VERSION : 0.1
   VAR_INPUT
      tcon_param : TCON_Param;
      send_buffer : "ADP.Message_Buffer.UDT";
   END_VAR
   VAR_IN_OUT
      requests : "Connection_Requests.UDT";
      saved_status : "Connection_Status.UDT";
   END_VAR
   VAR
      timers : "Connection_Status_Timers.UDT";
      TSEND : TSEND;
   END_VAR
   VAR_TEMP
      block_staus : "Connection_Status.UDT";
   END_VAR
BEGIN
   #TSEND(REQ := #requests.send,
          ID := #tcon_param.ID,
          DONE => #block_staus.done,
          BUSY => #block_staus.busy,
          ERROR => #block_staus.error,
          STATUS => #block_staus.status,
          DATA := #send_buffer);
   #requests.send := FALSE;
   "Send_Status.to_Control_Element"(requests := #requests,
                                    block_status := #block_staus,
                                    saved_status := #saved_status,
                                    timers := #timers);
END_FUNCTION_BLOCK

// folder: tcpip_connection/send/send_status

FUNCTION "Send_Status.Done" : Void   // FC168, SCL
{ S7_Optimized_Access := 'TRUE' }
VERSION : 0.1
   VAR_INPUT
      requests : "Connection_Requests.UDT";
      block_status : "Connection_Status.UDT";
   END_VAR
   VAR_IN_OUT
      saved_status : "Connection_Status.UDT";
   END_VAR
BEGIN
   "Send_Status.Set_Done"(block_status := #block_status,
                                requests := #requests,
                                saved_status := #saved_status);
   "Send_Status.Reset_Done"(block_status := #block_status,
                                  requests := #requests,
                                  saved_status := #saved_status);
END_FUNCTION

FUNCTION "Send_Status.Error" : Void   // FC169, SCL
{ S7_Optimized_Access := 'TRUE' }
VERSION : 0.1
   VAR_INPUT
      block_status : "Connection_Status.UDT";
      requests : "Connection_Requests.UDT";
   END_VAR
   VAR_IN_OUT
      off_delay : TOF_TIME;
      saved_status : "Connection_Status.UDT";
   END_VAR
BEGIN
   "Send_Status.Set_Error"(block_status := #block_status,
                                 requests := #requests,
                                 off_delay := #off_delay,
                                 saved_status := #saved_status);
END_FUNCTION

FUNCTION "Send_Status.Reset_Busy" : Void   // FC170, SCL
{ S7_Optimized_Access := 'TRUE' }
VERSION : 0.1
   VAR_INPUT
      requests : "Connection_Requests.UDT";
   END_VAR
   VAR_IN_OUT
      saved_status : "Connection_Status.UDT";
   END_VAR
BEGIN
   IF #requests.connect THEN
       #saved_status.busy := FALSE;
   END_IF;
END_FUNCTION

FUNCTION "Send_Status.Set_Busy" : Void   // FC171, SCL
{ S7_Optimized_Access := 'TRUE' }
VERSION : 0.1
   VAR_INPUT
      block_status : "Connection_Status.UDT";
      requests : "Connection_Requests.UDT";
   END_VAR
   VAR_IN_OUT
      off_delay : TOF_TIME;
      saved_status : "Connection_Status.UDT";
   END_VAR
   VAR_TEMP
      _et : Time;
   END_VAR
   VAR CONSTANT
      DELAY : Time := t#3s;
   END_VAR
BEGIN
   #off_delay(IN := #block_status.busy AND NOT #requests.disconnect,
              PT := #DELAY,
              Q => #saved_status.busy,
              ET => #_et);
END_FUNCTION

FUNCTION "Send_Status.Busy" : Void   // FC172, SCL
{ S7_Optimized_Access := 'TRUE' }
VERSION : 0.1
   VAR_INPUT
      block_status : "Connection_Status.UDT";
      requests : "Connection_Requests.UDT";
   END_VAR
   VAR_IN_OUT
      off_delay : TOF_TIME;
      saved_status : "Connection_Status.UDT";
   END_VAR
BEGIN
   "Send_Status.Set_Busy"(block_status := #block_status,
                                requests := #requests,
                                off_delay := #off_delay,
                                saved_status := #saved_status);
   "Send_Status.Reset_Busy"(requests := #requests,
                                  saved_status := #saved_status);
END_FUNCTION

FUNCTION "Send_Status.to_Control_Element" : Void   // FC173, SCL
{ S7_Optimized_Access := 'TRUE' }
VERSION : 0.1
   VAR_INPUT
      requests : "Connection_Requests.UDT";
      block_status : "Connection_Status.UDT";
   END_VAR
   VAR_IN_OUT
      saved_status : "Connection_Status.UDT";
      timers : "Connection_Status_Timers.UDT";
   END_VAR
BEGIN
   "Send_Status.Busy"(block_status := #block_status,
                            requests := #requests,
                            off_delay := #timers.busy,
                            saved_status := #saved_status);
   "Send_Status.Done"(requests := #requests,
                            block_status := #block_status,
                            saved_status := #saved_status);
   "Send_Status.Error"(block_status := #block_status,
                             requests := #requests,
                             off_delay := #timers.error,
                             saved_status := #saved_status);
   "Send_Status.Status"(block_status := #block_status,
                              requests := #requests,
                              saved_status := #saved_status,
                              status_timer := #timers.status);
END_FUNCTION

FUNCTION "Send_Status.Set_Done" : Void   // FC174, SCL
{ S7_Optimized_Access := 'TRUE' }
VERSION : 0.1
   VAR_INPUT
      block_status : "Connection_Status.UDT";
      requests : "Connection_Requests.UDT";
   END_VAR
   VAR_IN_OUT
      saved_status : "Connection_Status.UDT";
   END_VAR
BEGIN
   IF #block_status.done THEN
       #saved_status.done := TRUE;
   END_IF;
END_FUNCTION

FUNCTION "Send_Status.Reset_Done" : Void   // FC175, SCL
{ S7_Optimized_Access := 'TRUE' }
VERSION : 0.1
   VAR_INPUT
      block_status : "Connection_Status.UDT";
      requests : "Connection_Requests.UDT";
   END_VAR
   VAR_IN_OUT
      saved_status : "Connection_Status.UDT";
   END_VAR
BEGIN
   IF #requests.connect THEN
       #saved_status.done := FALSE;
   END_IF;
END_FUNCTION

FUNCTION "Send_Status.Set_Error" : Void   // FC176, SCL
{ S7_Optimized_Access := 'TRUE' }
VERSION : 0.1
   VAR_INPUT
      block_status : "Connection_Status.UDT";
      requests : "Connection_Requests.UDT";
   END_VAR
   VAR_IN_OUT
      off_delay : TOF_TIME;
      saved_status : "Connection_Status.UDT";
   END_VAR
   VAR_TEMP
      _et : Time;
   END_VAR
   VAR CONSTANT
      DELAY : Time := t#30s;
   END_VAR
BEGIN
   #off_delay(IN := #block_status.error,
              PT := #DELAY,
              Q => #saved_status.error,
              ET => #_et);
END_FUNCTION

FUNCTION "Send_Status.Save_Status" : Void   // FC177, SCL
{ S7_Optimized_Access := 'TRUE' }
VERSION : 0.1
   VAR_INPUT
      block_status : "Connection_Status.UDT";
   END_VAR
   VAR_IN_OUT
      saved_status : "Connection_Status.UDT";
      status_timer : TOF_TIME;
   END_VAR
   VAR_TEMP
      _delay_update : Bool;
      _et : Time;
   END_VAR
   VAR CONSTANT
      DELAY : Time := T#30S;
      IDLE : Word := 16#7000;
   END_VAR
BEGIN
   IF #block_status.status <> #IDLE THEN
       #saved_status.status := #block_status.status;
   END_IF;
   #status_timer(IN := #block_status.status <> #IDLE,
                 PT := #DELAY,
                 Q => #_delay_update,
                 ET => #_et);
   IF #_delay_update THEN
       RETURN;
   END_IF;
   #saved_status.status := #block_status.status;
END_FUNCTION

FUNCTION "Send_Status.Status" : Void   // FC178, SCL
{ S7_Optimized_Access := 'TRUE' }
VERSION : 0.1
   VAR_INPUT
      block_status : "Connection_Status.UDT";
      requests : "Connection_Requests.UDT";
   END_VAR
   VAR_IN_OUT
      saved_status : "Connection_Status.UDT";
      status_timer : TOF_TIME;
   END_VAR
BEGIN
   "Send_Status.Save_Status"(block_status := #block_status,
                                   saved_status := #saved_status,
                                   status_timer := #status_timer);
   "Send_Status.Clear_Status"(requests := #requests,
                                    saved_status := #saved_status);
END_FUNCTION

FUNCTION "Send_Status.Clear_Status" : Void   // FC179, SCL
{ S7_Optimized_Access := 'TRUE' }
VERSION : 0.1
   VAR_INPUT
      requests : "Connection_Requests.UDT";
   END_VAR
   VAR_IN_OUT
      saved_status : "Connection_Status.UDT";
   END_VAR
BEGIN
   IF #requests.connect THEN
       #saved_status.status := 0;
   END_IF;
END_FUNCTION

// folder: wire_hmi

FUNCTION "Wire_HMI.Input_Animations" : Void   // FC10, SCL
{ S7_Optimized_Access := 'TRUE' }
VERSION : 0.1
   VAR_IN_OUT
      wire : "Wire.HMI.UDT";
   END_VAR
BEGIN
   "Row_Data.Animate_In_Focus"(#wire.heat);
   "Row_Data.Animate_In_Focus"(#wire.carbon);
   "Row_Data.Animate_In_Focus"(#wire.calcium_silicon);
   "Row_Data.Animate_In_Focus"(#wire.aluminum);
   "Row_Data.Animate_In_Focus"(#wire.sulfur);
END_FUNCTION

FUNCTION "Wire_HMI.Initialize_Display" : Void   // FC29, SCL
{ S7_Optimized_Access := 'TRUE' }
VERSION : 0.1
   VAR_IN_OUT
      wire : "Wire.HMI.UDT";
   END_VAR
BEGIN
   "Screen_Background.Initialize"(#wire.background);
   "Row_Data.Initialize"(#wire.heat);
   "Row_Label.Initialize"(#wire.header);
   "Divider.Initialize"(#wire.divider);
   "Row_Data.Initialize"(#wire.carbon);
   "Row_Data.Initialize"(#wire.calcium_silicon);
   "Row_Data.Initialize"(#wire.aluminum);
   "Row_Data.Initialize"(#wire.sulfur);
   "Divider.Initialize"(#wire.bottom_border);
   "Divider.Hide_Line"(#wire.bottom_border);
END_FUNCTION

// folder: wire_message

FUNCTION_BLOCK "Wire_Message.Reset_Display_Driver"   // FB15, SCL
{ S7_Optimized_Access := 'TRUE' }
VERSION : 0.1
   VAR_INPUT
      send_buffer : "ADP.Message_Buffer.UDT";
   END_VAR
   VAR_IN_OUT
      interface : "Wire.HMI.UDT";
   END_VAR
   VAR
      "Message.Detect_Change" : "Message.Detect_Change";
      Reset_Display_Timer : TOF_TIME;
      old : Struct
         reset : Bool;
      END_STRUCT;
   END_VAR
   VAR_TEMP
      _message_changed : Bool;
      _et : Time;
      _reset_display : Bool;
   END_VAR
   VAR CONSTANT
      RESET_TIME : Time := T#10m;
   END_VAR
BEGIN
   #"Message.Detect_Change"(send_buffer := #send_buffer,
                            detected := #_message_changed);
   #Reset_Display_Timer(IN := #_message_changed,
                        PT := #RESET_TIME,
                        Q => #_reset_display,
                        ET => #_et);
   IF NOT #_reset_display AND #old.reset THEN
       "Wire_Message.Reset_Display"(#interface);
   END_IF;
   #old.reset := #_reset_display;
END_FUNCTION_BLOCK

FUNCTION_BLOCK "Wire_Message"   // FB25, SCL
{ S7_Optimized_Access := 'TRUE' }
VERSION : 0.1
   VAR_INPUT
      adp_liberary : "ADP.Encoded.UDT";
   END_VAR
   VAR_IN_OUT
      hmi_interface : "HMI_Interface.UDT";
      led_interface : "LED_Interface.UDT";
   END_VAR
   VAR
      mode : String;
      old : Struct
         mode : String;
      END_STRUCT;
      set_mode : "Wire_Message.Set_Mode";
      send_request : "Message.Request_Send";
      "Wire_Message.Reset_Display_Driver" : "Wire_Message.Reset_Display_Driver";
   END_VAR
BEGIN
   #set_mode(manual_request := #hmi_interface.connection_controls.wire.send.operation_button_actuate,
             mode := #mode);

   IF #mode = "AUTOMATIC" THEN
       #"Wire_Message.Reset_Display_Driver"(send_buffer := #led_interface.send_buffer,
                                            interface := #hmi_interface.wires);

       "Wire_Message.Assemble_Automatic_Message"(adp_library := #adp_liberary,
                                                 interface := #hmi_interface.wires,
                                                 send_buffer := #led_interface.send_buffer);
   END_IF;

   IF #mode = "MANUAL" AND #mode <> #old.mode THEN
       "Wire_Message.Assemble_Manual_Message"(adp_library := #adp_liberary,
                                              send_buffer := #led_interface.send_buffer);
   END_IF;

   #old.mode := #mode;

   #send_request(manual_request := #hmi_interface.connection_controls.wire.send.operation_button_actuate,
                 send_buffer := #led_interface.send_buffer,
                 send_request := #led_interface.requests.send);
END_FUNCTION_BLOCK

FUNCTION_BLOCK "Wire_Message.Set_Mode"   // FB27, SCL
{ S7_Optimized_Access := 'TRUE' }
VERSION : 0.1
   VAR_INPUT
      manual_request : Bool;
      automatic_request : Bool;
   END_VAR
   VAR_IN_OUT
      mode : String;
   END_VAR
   VAR
      manual_delay : TOF_TIME;
      old : Struct
         in_manual_delay : Bool;
      END_STRUCT;
   END_VAR
   VAR_TEMP
      _in_manual_delay : Bool;
      _et : Time;
   END_VAR
   VAR CONSTANT
      DELAY : Time := T#15S;
   END_VAR
BEGIN
   #manual_delay(IN := #manual_request AND NOT #manual_delay.Q,
                 PT := #DELAY,
                 Q => #_in_manual_delay,
                 ET => #_et);

   IF NOT #_in_manual_delay THEN
       #mode := "AUTOMATIC";
       #old.in_manual_delay := #_in_manual_delay;
       RETURN;
   END_IF;

   #mode := "MANUAL";
   #old.in_manual_delay := #_in_manual_delay;
   RETURN;
END_FUNCTION_BLOCK

FUNCTION "Wire_Message.Assemble_Automatic_Message" : Void   // FC180, SCL
{ S7_Optimized_Access := 'TRUE' }
VERSION : 0.1
   VAR_INPUT
      adp_library : "ADP.Encoded.UDT";
      interface : "Wire.HMI.UDT";
   END_VAR
   VAR_IN_OUT
      send_buffer : "ADP.Message_Buffer.UDT";
   END_VAR
   VAR_TEMP
      _count : UInt;
      _i : Int;
      _message : String;
      _rows : Array[0..5] of String;
      _send_buffer : "ADP.Message_Buffer.UDT";
   END_VAR
BEGIN
   REGION "MESSAGE HEADER"
       #_message := CONCAT_STRING(IN1 := #adp_library.file_system."00 Start of Header",
                                  IN2 := #adp_library.file_system."01 Address",
                                  IN3 := #adp_library.file_system."02 Start of Text",
                                  IN4 := #adp_library.file_system."03 Command & File",
                                  IN5 := #adp_library.formatting.size_and_face.normal_7);
   END_REGION


   REGION "TABLE ROWS"
       #_rows[0] := "Message.Assemble_Row"(adp_library := #adp_library,
                                           cell_0_value := 'HEAT',
                                           cell_0_color := #adp_library.formatting.color.yellow,
                                           cell_1_value := #interface.heat.cell_1_value,
                                           cell_1_color := '');

       #_rows[1] := "Message.Assemble_Row"(adp_library := #adp_library,
                                           cell_0_value := 'WIRE',
                                           cell_0_color := #adp_library.formatting.color.blue,
                                           cell_1_value := 'FEET',
                                           cell_1_color := '');


       #_rows[2] := "Message.Assemble_Row"(adp_library := #adp_library,
                                           cell_0_value := 'CARBON',
                                           cell_0_color := #adp_library.formatting.color.white,
                                           cell_1_value := #interface.carbon.cell_1_value,
                                           cell_1_color := '');

       #_rows[3] := "Message.Assemble_Row"(adp_library := #adp_library,
                                           cell_0_value := 'CAL/SIL',
                                           cell_0_color := '',
                                           cell_1_value := #interface.calcium_silicon.cell_1_value,
                                           cell_1_color := '');

       #_rows[4] := "Message.Assemble_Row"(adp_library := #adp_library,
                                           cell_0_value := 'ALUMINUM',
                                           cell_0_color := '',
                                           cell_1_value := #interface.aluminum.cell_1_value,
                                           cell_1_color := '');

       #_rows[5] := "Message.Assemble_Row"(adp_library := #adp_library,
                                           cell_0_value := 'SULFUR',
                                           cell_0_color := '',
                                           cell_1_value := #interface.sulfur.cell_1_value,
                                           cell_1_color := '');
       #_rows[5] := "String.Drop_Last_Character"(#_rows[5]);
   END_REGION


   REGION "CONCAT HEADER AND ROWS"
       FOR #_i := 0 TO 5 DO
           #_message := CONCAT_STRING(IN1 := #_message, IN2 := #_rows[#_i]);
       END_FOR;
   END_REGION


   REGION "END OF MESSAGE"
       #_message := CONCAT_STRING(IN1 := #_message, IN2 := #adp_library.file_system."04 END");
   END_REGION


   REGION "RETURN"
       Strg_TO_Chars(Strg := #_message,
                     pChars := 0,
                     Cnt => #_count,
                     Chars := #send_buffer.me);
   END_REGION
END_FUNCTION

FUNCTION "Wire_Message.Assemble_Manual_Message" : Void   // FC183, SCL
{ S7_Optimized_Access := 'TRUE' }
VERSION : 0.1
   VAR_INPUT
      adp_library : "ADP.Encoded.UDT";
   END_VAR
   VAR_IN_OUT
      send_buffer : "ADP.Message_Buffer.UDT";
   END_VAR
   VAR_TEMP
      _count : UInt;
      _i : Int;
      _message : String;
      _rows : Array[0..8] of String;
      _send_buffer : "ADP.Message_Buffer.UDT";
   END_VAR
BEGIN
   #_message := CONCAT_STRING(IN1 := #adp_library.file_system."00 Start of Header",
                              IN2 := #adp_library.file_system."01 Address",
                              IN3 := #adp_library.file_system."02 Start of Text",
                              IN4 := #adp_library.file_system."03 Command & File",
                              IN5 := 'WIRE COMMUNICATIONS TEST',
                              IN6 := #adp_library.file_system."04 END");


   Strg_TO_Chars(Strg := #_message,
                 pChars := 0,
                 Cnt => #_count,
                 Chars := #send_buffer.me);
END_FUNCTION

FUNCTION "Wire_Message.Reset_Display" : Void   // FC196, SCL
{ S7_Optimized_Access := 'TRUE' }
VERSION : 0.1
   VAR_IN_OUT
      interface : "Wire.HMI.UDT";
   END_VAR
   VAR CONSTANT
      BLANK : String;
   END_VAR
BEGIN
   #interface.heat.cell_1_value := #BLANK;
   #interface.carbon.cell_1_value := #BLANK;
   #interface.calcium_silicon.cell_1_value := #BLANK;
   #interface.aluminum.cell_1_value := #BLANK;
   #interface.sulfur.cell_1_value := #BLANK;
END_FUNCTION

// folder: wire_sign

FUNCTION "Wire_Sign.Set_Connection_Parameters" : Void   // FC128, SCL
{ S7_Optimized_Access := 'TRUE' }
VERSION : 0.1
   VAR_INPUT
      mode : String;
   END_VAR
   VAR_IN_OUT
      interface : "Connection_Parameters_HMI_Interface.UDT";
      saved : "Connection_Parameters.UDT";
   END_VAR
BEGIN
   IF #mode <> "WIRE" THEN
       RETURN;
   END_IF;
   "Connection_Parameters.Set_Parameters"(interface := #interface,
                                          saved :=#saved);
   RETURN;
END_FUNCTION

// folder: word

FUNCTION "Word.to_String" : String   // FC118, SCL
{ S7_Optimized_Access := 'TRUE' }
VERSION : 0.1
   VAR_INPUT
      value : Word;
   END_VAR
   VAR_TEMP
      _ret : String;
   END_VAR
BEGIN
   #"Word.to_String" := CONCAT_STRING(IN1 := "Byte.to_String"(#value.%B1),
                                      IN2 := "Byte.to_String"(#value.%B0));
END_FUNCTION

// folder: wstring

FUNCTION "WString.Split_Single" : Void   // FC15, SCL
{ S7_Optimized_Access := 'TRUE' }
VERSION : 0.1
   VAR_INPUT
      wstring_in : WString;
      delimeter : WString;
      pointer : Int;
   END_VAR
   VAR_IN_OUT
      sub_strings : Array[*] of WString;
   END_VAR
   VAR_TEMP
      _split : WString;
      _position : Int;
      _return : WString;
   END_VAR
BEGIN
   REGION "GET POSITION OF DELIMETER IN STRING"
       #_position := FIND(IN1 := #wstring_in,
                          IN2 := #delimeter);
   END_REGION

   REGION "BASE CASE"
       IF #_position = 0 THEN
           #sub_strings[#pointer] := #wstring_in;
           RETURN;
       END_IF;
   END_REGION


   REGION "RECURSIVE CASE"
       #sub_strings[#pointer] := LEFT(IN := #wstring_in, L := #_position - 1);
       "WString.Split_Single"(wstring_in := RIGHT(IN := #wstring_in, L := LEN(#wstring_in) - #_position),
                              delimeter := #delimeter,
                              "pointer" := #pointer + 1,
                              sub_strings := #sub_strings);
   END_REGION
END_FUNCTION

FUNCTION "WString.Find_Multiple.Breadth" : Int   // FC17, SCL
{ S7_Optimized_Access := 'TRUE' }
VERSION : 0.1
   VAR_INPUT
      body : WString;
      terms : Array[*] of WString[1];
   END_VAR
   VAR_TEMP
      _i : Int;
      _length : UDInt;
      _min : Int;
      _position : Int;
   END_VAR
   VAR CONSTANT
      BLANK : WString;
   END_VAR
BEGIN
   (* 
       Depth first search of 'body' for first occurance of any element of 'terms'.
       For depth first search use WString.Find_Multiple.Depth.
       Returns character postion in the string (1 indexed).
       E.G.: 
           - body := WSTRING#'today?'
           - terms := <WSTRING#>['?', 'ay']
           - returns --> 6
       E.G.:
           - body := WSTRING#'today?'
           - terms := <WSTRING#>['ay', '?']
           - returns --> 4
   *)

   #_length := "Any.Array.Length"(#terms);

   IF #_length = 0 OR #body = #BLANK THEN
       #"WString.Find_Multiple.Breadth" := 0;
       RETURN;
   END_IF;

   FOR #_i := 0 TO UDINT_TO_INT(#_length) - 1 DO
       #_position := FIND(IN1 := #body,
                          IN2 := #terms[#_i]);
       IF #_position = 0 THEN
           CONTINUE;
       END_IF;
       IF #_position < #_min OR #_min = 0 THEN
           #_min := #_position;
       END_IF;
   END_FOR;

   #"WString.Find_Multiple.Breadth" := #_min;
END_FUNCTION

FUNCTION "WString.Split_Multiple.Clean_Output" : Void   // FC25, SCL
{ S7_Optimized_Access := 'TRUE' }
VERSION : 0.1
   VAR_INPUT
      pointer : Int;
   END_VAR
   VAR_IN_OUT
      substrings : Array[*] of WString[20];
   END_VAR
   VAR_TEMP
      _i : Int;
   END_VAR
   VAR CONSTANT
      BLANK : WString;
   END_VAR
BEGIN
   FOR #_i := #"pointer" TO UDINT_TO_INT("Any.Array.Length"(#substrings)) - 1 DO
       #substrings[#_i] := wstring#'';
   END_FOR;
END_FUNCTION

FUNCTION "WString.Split_Multiple" : Void   // FC36, SCL
{ S7_Optimized_Access := 'TRUE' }
VERSION : 0.1
   VAR_INPUT
      wstring_in : WString;
      delimeters : Array[*] of WString[1];
      pointer : Int;
   END_VAR
   VAR_OUTPUT
      substrings : Array[*] of WString[20];
   END_VAR
   VAR_TEMP
      _i : Int;
      _position : Int;
      _return : WString;
      _split : WString;
   END_VAR
BEGIN
   REGION "GET POSITION OF DELIMETER IN STRING"
       #_position := "WString.Find_Multiple.Breadth"(body := #wstring_in,
                                                     terms := #delimeters);
   END_REGION

   REGION "BASE CASE"
       IF #_position = 0 THEN
           #substrings[#pointer] := #wstring_in;
           "WString.Split_Multiple.Clean_Output"("pointer" := #pointer + 1,
                                                 substrings := #substrings);
           RETURN;
       END_IF;
   END_REGION


   REGION "RECURSIVE CASE"
       #substrings[#pointer] := LEFT(IN := #wstring_in, L := #_position);
       "WString.Split_Multiple"(wstring_in := RIGHT(IN := #wstring_in, L := LEN(#wstring_in) - #_position),
                                delimeters := #delimeters,
                                "pointer" := #pointer + 1,
                                substrings => #substrings);
   END_REGION
END_FUNCTION

FUNCTION "WString.Search_Array" : Int   // FC67, SCL
{ S7_Optimized_Access := 'TRUE' }
VERSION : 0.1
   VAR_INPUT
      "array" : Array[*] of WString;
      search_term : WString;
   END_VAR
   VAR_TEMP
      _i : Int;
      _length : Int;
   END_VAR
BEGIN
   REGION "SEARCH ARRAY"    
       #_length := UDINT_TO_INT("Any.Array.Length"(#array)) - 1;
       FOR #_i := 0 TO #_length DO
           IF #array[#_i] = #search_term THEN
               #"WString.Search_Array" := #_i;
               RETURN;
           END_IF;
       END_FOR;
   END_REGION

   REGION "RETURN"
       #"WString.Search_Array" := "NULL_TOKEN";
       RETURN;
   END_REGION
END_FUNCTION

FUNCTION "WString.Reverse_Array" : Void   // FC68, SCL
{ S7_Optimized_Access := 'TRUE' }
VERSION : 0.1
   VAR_INPUT
      null_token : WString;
   END_VAR
   VAR_IN_OUT
      wstring_array : Array[*] of WString;
   END_VAR
   VAR_TEMP
      _has_data_count : Int;
      _i : Int;
      _p_swap : Int;
      _temp : WString;
   END_VAR
   VAR CONSTANT
      NOT_FOUND : Int := -1;
   END_VAR
BEGIN
   REGION "CHECK FOR FIRST EMPTY POSITION"
       #_has_data_count := "WString.Search_Array"(array := #wstring_array,
                                                  search_term := #null_token);
   END_REGION


   REGION "EXIT ON EMPTY ARRAY"
       IF #_has_data_count = 0 THEN
           RETURN;
       END_IF;
   END_REGION


   REGION "ARRAY IS FULL"
       IF #_has_data_count = #NOT_FOUND THEN
           #_has_data_count := UDINT_TO_INT("Any.Array.Length"(#wstring_array));
       END_IF;
   END_REGION


   REGION "ADJUST TO ZERO INDEX"
       #_has_data_count -= 1;
   END_REGION


   REGION "SWAP ELEMENTS"
       FOR #_i := 0 TO #_has_data_count / 2 DO
           #_p_swap := #_has_data_count - #_i;
           #_temp := #wstring_array[#_i];
           #wstring_array[#_i] := #wstring_array[#_p_swap];
           #wstring_array[#_p_swap] := #_temp;
       END_FOR;
   END_REGION


   REGION "DONE"
       RETURN;
   END_REGION
END_FUNCTION

// ===== library types =====

TYPE "Row.UDT"
   STRUCT
      background_animate : DInt;
      background_visible : Bool;
      cell_0_animate : DInt;
      cell_0_visible : Bool;
      cell_1_active : Bool;
      cell_1_animate : DInt;
      cell_1_enable : Bool;
      cell_1_input_finished : Bool;
      cell_1_value : String[50];
      cell_1_visible : Bool;
   END_STRUCT;
END_TYPE

TYPE "Navigation.UDT"
   STRUCT
      background_animate : DInt;
      background_visible : Bool;
      bottom_line_animate : DInt;
      bottom_line_visible : Bool;
      communications_status_actuate : Bool;
      communications_status_animate : DInt;
      communications_status_cover_animate : DInt;
      communications_status_cover_visible : Bool;
      communications_status_enable : Bool;
      communications_status_visible : Bool;
      material_actuate : Bool;
      material_animate : DInt;
      material_cover_animate : DInt;
      material_cover_visible : Bool;
      material_enable : Bool;
      material_visible : Bool;
      wire_actuate : Bool;
      wire_animate : DInt;
      wire_cover_animate : DInt;
      wire_cover_visible : Bool;
      wire_enable : Bool;
      wire_visible : Bool;
   END_STRUCT;
END_TYPE

// folder: connection

TYPE "Connection_Parameters_HMI.UDT"
   STRUCT
      back_actuate : Bool;
      back_animate : DInt;
      back_enable : Bool;
      back_visible : Bool;
      header_animate : DInt;
      header_value : String[25];
      header_visible : Bool;
      id_label_animate : DInt;
      id_label_visible : Bool;
      id_entry_active : Bool;
      id_entry_animate : DInt;
      id_entry_input_finished : Bool;
      id_entry_enable : Bool;
      id_entry_value : String[6];
      id_entry_visible : Bool;
      ip_address_label_animate : DInt;
      ip_address_label_visible : Bool;
      ip_address_entry_active : Bool;
      ip_address_entry_animate : DInt;
      ip_address_entry_enable : Bool;
      ip_address_entry_input_finished : Bool;
      ip_address_entry_value : String[15];
      ip_address_entry_visible : Bool;
      port_label_animate : DInt;
      port_label_visible : Bool;
      port_entry_active : Bool;
      port_entry_animate : DInt;
      port_entry_enable : Bool;
      port_entry_input_finished : Bool;
      port_entry_value : String[6];
      port_entry_visible : Bool;
   END_STRUCT;
END_TYPE

// folder: connection_detail

TYPE "Connection_Status_Detail.HMI.UDT"
   STRUCT
      back_button_actuate : Bool;
      back_button_enable : Bool;
      back_button_visible : Bool;
      detailed_status_animate : DInt;
      detailed_status_visible : Bool;
      detailed_status_list_selector : DInt;
      detailed_status_message_selector : DInt;
      display_payload_button_actuate : Bool;
      display_payload_button_animate : DInt;
      display_payload_button_enable : Bool;
      display_payload_button_visible : Bool;
      header_animate : DInt;
      header_selector : DInt;
      header_visible : Bool;
      payload_animate : DInt;
      payload_text : String;
      payload_visible : Bool;
   END_STRUCT;
END_TYPE

// folder: (top level)

FUNCTION "Array.Any.Length" : UDInt   // FC16, SCL
{ S7_Optimized_Access := 'TRUE' }
VERSION : 0.1
   VAR_INPUT
      "array" : Variant;
   END_VAR
   VAR_TEMP
      status : DInt;
      ret : UDInt;
   END_VAR
BEGIN
   #ret := CountOfElements(#array);
   #"Array.Any.Length" := #ret;
END_FUNCTION

// folder: color

FUNCTION "Color.Decode_String" : DInt   // FC14, SCL
{ S7_Optimized_Access := 'TRUE' }
VERSION : 0.1
   VAR_INPUT
      color : String;   // enter rgb value with comma, semicolon, or underscore as delimeter. e.g.: '200,100,200' or '195_168_0'
   END_VAR
   VAR_TEMP
      _delimeters : Array[0..2] of String[1];
      _substrings : Array[0..2] of String[20];
      _red : DInt;
      _green : DInt;
      _blue : DInt;
   END_VAR
BEGIN
   #_delimeters[0] := ',';
   #_delimeters[1] := ';';
   #_delimeters[2] := '_';
   "String.Split_Multiple"(string_in:=#color,
                           delimeters:=#_delimeters,
                           "pointer":=0,
                           substrings=>#_substrings);
   #_red := STRING_TO_DINT(#_substrings[0]) * 1_000_000;
   #_green := STRING_TO_DINT(#_substrings[1]) * 1_000;
   #_blue := STRING_TO_DINT(#_substrings[2]);
   #"Color.Decode_String" := #_red + #_green + #_blue;
END_FUNCTION

// ===== library: MasterCopy "Copy of PLC data types in ADP Data" =====

// folder: ADP Data

TYPE "ADP: Encoded"
VERSION : 0.1
   STRUCT
      file_system : "ADP: Encoded: File System";
      formatting : "ADP: Encoded: Formatting";
   END_STRUCT;
END_TYPE

TYPE "ADP: Decoded"
   STRUCT
      color : "ADP: Decoded: Color";
      flash : "ADP: Decoded: Flash";
      horizontal_alignment : "ADP: Decoded: Horizontal Alignment";
      line_control : "ADP: Decoded: Line Control";
      scroll_speed : "ADP: Decoded: Scroll Speed";
      size_and_face : "ADP: Decoded: Size and Face";
      vertical_alignment : "ADP: Decoded: Vertical Alignment";
   END_STRUCT;
END_TYPE

TYPE "ADP: Decoded: Color"
   STRUCT
      black : String[8] := 'black';
      blue : String[8] := 'blue';
      green : String[8] := 'green';
      mix_1 : String[8] := 'mix 1';
      mix_2 : String[8] := 'mix 2';
      mix_3 : String[8] := 'mix 3';
      mix_4 : String[8] := 'mix 4';
      red : String[8] := 'red';
      white : String[8] := 'white';
      yellow : String[8] := 'yellow';
   END_STRUCT;
END_TYPE

TYPE "ADP: Decoded: Flash"
   STRUCT
      off : String[8] := 'off';
      on : String[8] := 'on';
   END_STRUCT;
END_TYPE

TYPE "ADP: Decoded: Horizontal Alignment"
   STRUCT
      center : String[8] := 'center';
      left : String[8] := 'left';
      right : String[8] := 'right';
   END_STRUCT;
END_TYPE

TYPE "ADP: Message Formats: Encoded"
   STRUCT
      color : String [5];
      flash : String [5];
      scroll_speed : String [5];
      size_and_face : String [5];
      vertical_alignment : String [5];
      horizontal_alignment : String [5];
   END_STRUCT;
END_TYPE

TYPE "ADP: Message Formats: Decoded"
   STRUCT
      color : String [20];
      flash : String [20];
      scroll_speed : String [20];
      size_and_face : String [20];
      vertical_alignment : String [20];
      horizontal_alignment : String [20];
   END_STRUCT;
END_TYPE

TYPE "ADP: Decoded: Scroll Speed"
   STRUCT
      slowest : String[9] := 'slowest';
      slow : String[9] := 'slow';
      normal : String[9] := 'normal';
      fast : String[9] := 'fast';
      fastest : String[9] := 'fastest';
   END_STRUCT;
END_TYPE

TYPE "ADP: Decoded: Size and Face"
   STRUCT
      bold_5 : String[11] := 'bold 5';
      bold_11 : String[11] := 'bold 11';
      bold_14 : String[11] := 'bold 14';
      bold_15 : String[11] := 'bold 15';
      bold_16 : String[11] := 'bold 16';
      bold_22 : String[11] := 'bold 22';
      bold_30 : String[11] := 'bold 30';
      bold_32 : String[11] := 'bold 32';
      bold_40 : String[11] := 'bold 40';
      normal_5 : String[11] := 'normal 5';
      normal_7 : String[11] := 'normal 7';
      normal_9 : String[11] := 'normal 9';
      normal_11 : String[11] := 'normal 11';
      normal_14 : String[11] := 'normal 14';
      normal_15 : String[11] := 'normal 15';
      normal_16 : String[11] := 'normal 16';
      normal_22 : String[11] := 'normal 22';
      normal_24 : String[11] := 'normal 24';
      normal_30 : String[11] := 'normal 30';
      normal_32 : String[11] := 'normal 32';
      normal_40 : String[11] := 'normal 40';
   END_STRUCT;
END_TYPE

TYPE "ADP: Decoded: Vertical Alignment"
   STRUCT
      bottom_hold : String[15] := 'bottom hold';
      fill_hold : String[15] := 'fill hold';
      middle_hold : String[15] := 'middle hold';
      top_hold : String[15] := 'top hold';
      bottom_scroll : String[15] := 'bottom scroll';
      fill_scroll : String[15] := 'fill scroll';
      middle_scroll : String[15] := 'middle scroll';
      top_scroll : String[15] := 'top scroll';
   END_STRUCT;
END_TYPE

TYPE "ADP: Encoded: File System"
   STRUCT
      "00 Start of Header" : String[5] := '$01';
      "01 Address" : String[5] := 'Z00';
      "02 Start of Text" : String[5] := '$02';
      "03 Command & File" : String[5] := 'AA';
      "04 END" : String[5] := '$04';
   END_STRUCT;
END_TYPE

TYPE "ADP: Encoded: Formatting"
   STRUCT
      color : "ADP: Encoded: Formatting: Color";
      flashing : "ADP: Encoded: Formatting: Flashing";
      horizontal_alignment : "ADP: Encoded: Formatting: Horizontal Alignment";
      line_control : "ADP: Encoded: Formatting: Line Control";
      scroll_speed : "ADP: Encoded: Formatting: Scroll Speed";
      size_and_face : "ADP: Encoded: Formatting: Size and Face";
      vertical_alignment : "ADP: Encoded: Formatting: Vertical Alignment";
   END_STRUCT;
END_TYPE

TYPE "ADP: Encoded: Formatting: Color"
   STRUCT
      black : String[5] := '$1C0';
      blue : String[5] := '$1C8';
      green : String[5] := '$1C2';
      mix_1 : String[5] := '$1C4';
      mix_2 : String[5] := '$1C5';
      mix_3 : String[5] := '$1C6';
      mix_4 : String[5] := '$1CY';
      red : String[5] := '$1C1';
      white : String[5] := '$1C9';
      yellow : String[5] := '$1C3';
   END_STRUCT;
END_TYPE

TYPE "ADP: Encoded: Formatting: Flashing"
   STRUCT
      off : String[5] := '$070';
      on : String[5] := '$071';
   END_STRUCT;
END_TYPE

TYPE "ADP: Encoded: Formatting: Size and Face"
   STRUCT
      bold_5 : String[5] := '$1AG';
      bold_11 : String[5] := '$1AH';
      bold_14 : String[5] := '$1A5';
      bold_15 : String[5] := '$1A6';
      bold_16 : String[5] := '$1A7';
      bold_22 : String[5] := '$1AC';
      bold_30 : String[5] := '$1AI';
      bold_32 : String[5] := '$1AJ';
      bold_40 : String[5] := '$1AK';
      normal_5 : String[5] := '$1A0';
      normal_7 : String[5] := '$1A1';
      normal_9 : String[5] := '$1A8';
      normal_11 : String[5] := '$1A9';
      normal_14 : String[5] := '$1A2';
      normal_15 : String[5] := '$1A3';
      normal_16 : String[5] := '$1A4';
      normal_22 : String[5] := '$1AA';
      normal_24 : String[5] := '$1AB';
      normal_30 : String[5] := '$1AD';
      normal_32 : String[5] := '$1AE';
      normal_40 : String[5] := '$1AF';
   END_STRUCT;
END_TYPE

TYPE "ADP: Encoded: Formatting: Horizontal Alignment"
   STRUCT
      center : String[5] := '$L1';
      left : String[5] := '$L0';
      right : String[5] := '$L2';
   END_STRUCT;
END_TYPE

TYPE "ADP: Encoded: Formatting: Vertical Alignment"
   STRUCT
      middle_hold : String[5] := '$1B b';
      fill_hold : String[5] := '$1B"b';
      bottom_hold : String[5] := '$1B&b';
      top_hold : String[5] := '$1B0b';
      bottom_scroll : String[5] := '$1B a';
      fill_scroll : String[5] := '$1B"a';
      middle_scroll : String[5] := '$1B&a';
      top_scroll : String[5] := '$1B0a';
   END_STRUCT;
END_TYPE

TYPE "ADP: Encoded: Formatting: Scroll Speed"
   STRUCT
      slowest : String[5] := '$15';
      slow : String[5] := '$16';
      normal : String[5] := '$17';
      fast : String[5] := '$18';
      fastest : String[5] := '$19';
   END_STRUCT;
END_TYPE

TYPE "ADP: Encoded: Formatting: Line Control"
   STRUCT
      new_line : String[5] := '$R';
      word_wrap : String[5] := '';
   END_STRUCT;
END_TYPE

TYPE "ADP: Decoded: Line Control"
   STRUCT
      new_line : String[9] := 'new line';
      word_wrap : String[9] := 'word wrap';
   END_STRUCT;
END_TYPE

(* ===== HMI "HMI_RT_1" =====
system functions are stored by id; their names below are inferred from use
connection "HMI_Connection_1": ETHERNET, S7_1200_OMS

HMI tags "Default tag table"
   "Clock_Byte" : Byte = PLC Clock_Byte AT %MB0, 100 ms
   "HMI_Interface.Data_materials" : Materials.HMI.UDT = PLC "HMI_Interface.Data".materials AT %DB1.DBB0, 100 ms
   "HMI_Interface.Data_navigation" : Navigation.HMI.UDT = PLC "HMI_Interface.Data".navigation AT %DB1.DBW0, 100 ms
   "HMI_Interface.Data_wires" : Wire.HMI.UDT = PLC "HMI_Interface.Data".wires AT %DB1.DBW0, 100 ms
   "HMI_Interface.Data_meta" : HMI_Meta.UDT = PLC "HMI_Interface.Data".meta AT %DB1.DBW0, 100 ms
   "HMI_Interface.Data_connection_controls" : Connection_Status.HMI.UDT = PLC "HMI_Interface.Data".connection_controls AT %DB1.DBW0, 100 ms
   "disconnect" : DInt AT %DB1.DBD0
   "connect" : DInt, internal
   "send" : DInt, internal
   "HMI_Interface.Data_connection_status_details" : Connection_Detail.HMI.UDT = PLC "HMI_Interface.Data".connection_status_details AT %DB1.DBW0, 100 ms
   "HMI_Interface.Data_connection_parameters" : Connection_Paramters_HMI.UDT = PLC "HMI_Interface.Data".connection_parameters, 100 ms

text list "Send Code Descriptions Long": 0 'Send job completed without error.'; 28672 'No job processing active.'; 28673 'Start of job execution, data is being sent. When processing this job, the operating system accesses the data in the DATA send area.'; 28674 'Job executing (REQ irrelevant). When processing this job, the operating system accesses the data in the DATA send area.'; 32901 'The LEN parameter is greater than the highest permitted value (65536). DATA and LEN parameters both have the value "0".'; 32902 'The ID parameter is outside the permitted address range (1..0xFFF).'; 32904 'The LEN parameter is greater than the area specified in DATA.'; 32929 'Communication error: The specified connection has not yet been established. The specified connection is being terminated. Transfer via thisconnection is not possible. The interface is being re-initialized.'; 32947 'The protocol variant (ConnectionType parameter in the connection description) is set to UDP. Use the instruction "TUSEND" with a UDP connection.'; 32963 'A block with this ID is already being processed in a different priority group. Internal lack of resources.'; 32964 'Temporary communication error: The connection cannot be established to the partner at this time. The interface is receiving new parameter settings or the connection is being established.'; 32965 'Connection terminated by the communication partner.'; 32966 'Network error. Communication partner cannot be reached.'; 32967 'Execution timeout'; 65535 'Function not yet called.'

text list "Connection Details Header": 0 'NO STATE'; 1 'DISCONNECTION STATUS'; 2 'CONNECTION STATUS'; 3 'SEND STATUS'

text list "Disconnect Code Descriptions Long": 0 'Connection terminated successfully.'; 28672 'No job processing active.'; 28673 'Start of job processing, connection being terminated.'; 28674 'Intermediate call (REQ irrelevant), connection being terminated.'; 32902 'The ID parameter is not in the permitted value range.'; 32931 'Attempt is being made to terminate a non-existent connection or the connection is already terminated.'; 32964 'Temporary communication error: New parameters are being assigned to the interface or the connection is currently being established.'; 65535 'In connect state.'

text list "Connect Code Descriptions Long": 0 'Connection successfully established.'; 28672 'No job processing active'; 28673 'Start job execution, establish connection.'; 28674 'Connection is being established (REQ irrelevant).'; 32901 'Connection ID (ID parameter) is already being used by a configured connection.'; 32902 'The ID parameter is outside the valid range.'; 32903 'Maximum number of connections reached; no additional connection possible'; 32905 'The CONNECT parameter does not point to a data block.'; 32922 'The structure at the CONNECT parameter is not supported on an integrated interface or the length is invalid or an incorrect "InterfaceID" is specified in the connection description (SDT).'; 32923 'The element InterfaceId within the TCON_xxx structure does not reference a hardware identifier of a CPU or CM/CP interface or has the value "0".'; 32928 'Group error for error codes W#16#80A1 and W#16#80A2.'; 32929 'The specified connection or the port is already being used.'; 32930 'Local or remote port is being used by the system.'; 32931 'Attempt being made to re-establish an existing connection.'; 32932 'IP address of the remote endpoint of the connection is invalid, in other words, it matches the IP address of the local partner.'; 32933 'Connection ID is already in use.'; 32935 'Communication error: You executed "TDISCON" before "TCON" had completed.'; 32946 'The CONNECT parameter points to a data block that was generated with the attribute "Only store in load memory".'; 32948 'ISO-on-TCP violation: local_tsap_id_len >= B#16#02 local_tsap_id[1] = B#16#E0 local_tsap_id_len >= B#16#03 local_tsap_id[1] is ASCII chr local_tsap_id[1] is ASCII cha and local_tsap_id_len >= B#16#03'; 32949 'Only passive connection establishment is permitted for connection type 13 = UDP.'; 32950 'Parameter assignment error at the connection_type parameter of the SDT TCON_Param.'; 32951 'Error in one of the following parameters of the data block for connection description: block_length, local_tsap_id_len, rem_subnet_id_len, rem_staddr_len, rem_tsap_id_len, next_staddr_len. Note: If you call TCON in TCP for the passive end, local_tsap_id_len must have the value 2 and rem_tsap_id_len the value 0.'; 32952 'Connection description of the structure element ID and the block parameter ID are not identical.'; 32963 'All connection resources are in use.'; 32964 'Temporary communication error: Firewall Pending Parameterization Pending Disconnect'; 65535 'In disconnect state.'; 32966 'The connection partner could not be reached.'

text list "Disconnect Code Descriptions Short": 0 'DISCONNECTION SUCCESSFUL'; 28672 'NO JOB'; 28673 'JOB STARTED'; 28674 'REQUEST DURING EXECUTION'; 32902 'ID INVALID: OUT OF RANGE'; 32931 'CONNECTION ALREADY TERMINATED'; 32964 'REQUEST DURING PARAM ASSIGNMENT'; 65535 'STATE: CONNECT'

text list "Send Code Descriptions Short": 0 'SEND SUCCESSFUL'; 28672 'NO JOB'; 28673 'DATA ACCESSED DURING JOB'; 28674 'JOB PROCESSING'; 32901 'MAX LENGTH EXCEEDED'; 32902 'INVALID ID OUT OF RANGE'; 32904 'LENGTH EXCEEDS DATA RANGE'; 32929 'NO CONNECTION'; 32947 'UDP CONNECTION'; 32963 'CONNECTION BUSY'; 32964 'REQUEST DURING PARAM ASSIGNMENT'; 32965 'PARTNER TERMINATED CONNECTION'; 32966 'PARTNER UNAVAILABLE'; 32967 'TIMEOUT'; 65535 'NOT CALLED'

text list "Connect Code Descriptions Short": 0 'CONNECTION SUCCESSFUL'; 28672 'NO JOB'; 28673 'START JOB'; 28674 'PROCESSING JOB'; 32901 'ID INVALID: ALREADY IN USE'; 32902 'ID INVALID: OUT OF RANGE'; 32903 'MAX CONNECTIONS REACHED'; 32905 'NO CONNECTION DATA STORED'; 32922 'INVALID CONNECTION DATA'; 32923 'NO CONNECTION HARDWARE'; 32928 'GROUP ERROR'; 32929 'LOCAL PORT IN USE'; 32930 'REMOTE PORT IN USE'; 32931 'CONNECTION ALREADY ESTABLISHED'; 32932 'INVALID IP ADDRESS'; 32933 'DUPLICATE CONNECTION ID'; 32935 'DICONNECT REQUEST WHILE CONNECTING'; 32946 'CONNECT DATA IN LOAD MEMORY'; 32948 'ISO ON TCP VIOLATION'; 32949 'NON PASSIVE UDP CONNECTION REQUEST'; 32950 'INVALID CONNECTION TYPE'; 32951 'CONNECTION PARAMETER ERROR'; 32952 'DATA/PARAMETER MISMATCH'; 32963 'MAX CONNECTIONS EXCEEDED'; 32964 'FIREWALL'; 65535 'STATE: DISCONNECT'; 32966 'PARTNER UNAVAILABLE'

Template "Navigation" 800x480
   ScreenModuleView "Navigation_1" at 0,0 size 800x65; ScreenModuleType ""
      Guid_{11997190-7796} <- "HMI_Interface.Data_navigation"
      on Guid_{11997190-7994}: ActivateScreen("02_Materials", 0)
      on Guid_{11997190-7997}: ActivateScreen("01_Wires", 0)
      on Guid_{11997190-23512}: ActivateScreen("03_Connection_Control", 0)

screen "01_Wires" 800x480, template "Navigation"
   on GenerateScreen: SetTag("screen_number", 1)
   ScreenModuleView "heat" at 100,75 size 600x65; Guid_{11997190-6447} 'HEAT'; ScreenModuleType ""
      Guid_{11997190-5401} <- "heat"
   ScreenModuleView "label" at 100,140 size 600x65; Guid_{11997190-7215} 'FEET'; ScreenModuleType ""
      Guid_{11997190-5401} <- "header"
   ScreenModuleView "divider" at 100,205 size 600x5; ScreenModuleType ""
      Guid_{11997190-7534} <- "divider"
   ScreenModuleView "carbon" at 100,210 size 600x65; Guid_{11997190-6447} 'CARBON'; ScreenModuleType ""
      Guid_{11997190-5401} <- "carbon"
   ScreenModuleView "calcium_silicon" at 100,275 size 600x65; Guid_{11997190-6447} 'CAL/SIL'; ScreenModuleType ""
      Guid_{11997190-5401} <- "calcium_silicon"
   ScreenModuleView "aluminium" at 100,340 size 600x65; Guid_{11997190-6447} 'ALUMINIUM'; ScreenModuleType ""
      Guid_{11997190-5401} <- "aluminum"
   ScreenModuleView "sulfur" at 100,405 size 600x65; Guid_{11997190-6447} 'SULFUR'; ScreenModuleType ""
      Guid_{11997190-5401} <- "sulfur"
   ScreenModuleView "bottom_border" at 100,470 size 600x5; ScreenModuleType ""
      Guid_{11997190-7534} <- "bottom_border"
   Rectangle "Rectangle_1" at 0,65 size 800x415
      Appearance <- "color"
      Visibility <- "visible"

screen "02_Materials" 800x480, template "Navigation"
   on GenerateScreen: SetTag("screen_number", 2)
   ScreenModuleView "heat" at 100,87 size 600x40; Guid_{11997190-6447} 'HEAT'; ScreenModuleType ""
      Guid_{11997190-5401} <- "heat"
   ScreenModuleView "material_label" at 100,127 size 600x40; ScreenModuleType ""
      Guid_{11997190-5401} <- "header"
   ScreenModuleView "divider" at 100,167 size 600x5; ScreenModuleType ""
      Guid_{11997190-7534} <- "divider"
   ScreenModuleView "manganese" at 100,172 size 600x40; Guid_{11997190-6447} 'MANGANESE'; ScreenModuleType ""
      Guid_{11997190-5401} <- "manganese"
   ScreenModuleView "silicon" at 100,212 size 600x40; Guid_{11997190-6447} 'SILICON'; ScreenModuleType ""
      Guid_{11997190-5401} <- "silicon"
   ScreenModuleView "chromium" at 100,252 size 600x40; Guid_{11997190-6447} 'CHROMIUM'; ScreenModuleType ""
      Guid_{11997190-5401} <- "chromium"
   ScreenModuleView "vanadium" at 100,292 size 600x40; Guid_{11997190-6447} 'VANADIUM'; ScreenModuleType ""
      Guid_{11997190-5401} <- "vanadium"
   ScreenModuleView "nickel" at 100,332 size 600x40; Guid_{11997190-6447} 'NICKEL'; ScreenModuleType ""
      Guid_{11997190-5401} <- "nickel"
   ScreenModuleView "molybdenum" at 100,372 size 600x40; Guid_{11997190-6447} 'MOLYBDENUM'; ScreenModuleType ""
      Guid_{11997190-5401} <- "molybdenum"
   ScreenModuleView "bottom_border" at 100,452 size 600x5; ScreenModuleType ""
      Guid_{11997190-7534} <- "bottom_border"
   ScreenModuleView "custom" at 100,412 size 600x40; ScreenModuleType ""
      Guid_{11997190-5401} <- "custom"
   Rectangle "screen_background" at 0,65 size 800x415
      Appearance <- "color"
      Visibility <- "visible"

screen "03_Connection_Control" 800x480, template "Navigation"
   on GenerateScreen: SetTag("screen_number", 3)
   Rectangle "screen_background" at 0,65 size 800x415
      Appearance <- "color"
      Visibility <- "visible"
   ScreenModuleView "wire_header" at 5,70 size 392x55; Guid_{11997190-22834} 'WIRE SIGN COMMUNICATIONS'; Guid_{11997190-31866} 'WIRE SIGN CONNECTION CONTROLS'; ScreenModuleType ""
      Guid_{11997190-22821} <- "header"
      on Guid_{11997190-31700}: ActivateScreen("05_Connection_Parameters", 0)
   ScreenModuleView "wire_disconnect" at 5,130 size 392x110; Guid_{11997190-22931} 'D'; ScreenModuleType ""
      Guid_{11997190-22837} <- "disconnect"
      Guid_{11997190-22858} <- "disconnect"
      on Guid_{11997190-23485}: ActivateScreen("04_Connection_Status_Details", 0)
   ScreenModuleView "wire_connect" at 5,245 size 392x110; Guid_{11997190-22931} 'C'; ScreenModuleType ""
      Guid_{11997190-22837} <- "connect"
      Guid_{11997190-22858} <- "connect"
      on Guid_{11997190-23485}: ActivateScreen("04_Connection_Status_Details", 0)
   ScreenModuleView "wire_send" at 5,360 size 392x110; ScreenModuleType ""
      Guid_{11997190-22837} <- "send"
      Guid_{11997190-22858} <- "send"
      on Guid_{11997190-23485}: ActivateScreen("04_Connection_Status_Details", 0)
   ScreenModuleView "material_header" at 403,70 size 392x55; Guid_{11997190-22834} 'MATERIAL SIGN COMMUNICATIONS'; Guid_{11997190-31866} 'MATERIAL SIGN CONNECTION CONTROLS'; ScreenModuleType ""
      Guid_{11997190-22821} <- "header"
      on Guid_{11997190-31700}: ActivateScreen("05_Connection_Parameters", 0)
   ScreenModuleView "material_disconnect" at 403,130 size 392x110; Guid_{11997190-22931} 'D'; ScreenModuleType ""
      Guid_{11997190-22837} <- "disconnect"
      Guid_{11997190-22858} <- "disconnect"
      on Guid_{11997190-23485}: ActivateScreen("04_Connection_Status_Details", 0)
   ScreenModuleView "material_connect" at 403,245 size 392x110; Guid_{11997190-22931} 'C'; ScreenModuleType ""
      Guid_{11997190-22837} <- "connect"
      Guid_{11997190-22858} <- "connect"
      on Guid_{11997190-23485}: ActivateScreen("04_Connection_Status_Details", 0)
   ScreenModuleView "material_send" at 403,360 size 392x110; ScreenModuleType ""
      Guid_{11997190-22837} <- "send"
      Guid_{11997190-22858} <- "send"
      on Guid_{11997190-23485}: ActivateScreen("04_Connection_Status_Details", 0)

screen "04_Connection_Status_Details" 800x480, template "Navigation"
   on GenerateScreen: SetTag("screen_number", 4)
   Rectangle "screen_background" at 0,65 size 800x415
      Visibility <- "visible"
      Appearance <- "color"
   ScreenModuleView "Communications_Details_1" at 5,70 size 790x405; ScreenModuleType ""
      Guid_{11997190-25821} <- "HMI_Interface.Data_connection_status_details"
      on Guid_{11997190-25792}: ActivateScreen("03_Connection_Control", 0)

